(* Logix 5000 project; controller PLC_MCC1201_220AP1 vendor 1 type 14 code 164 rev 35.11; software revision 35.00 *) (continued)
   OSR_xStopCycle : BOOL;   // OSR stop cycle
   OS_xAreaSafetyOK : BOOL;   // OS area safety ok
   OS_xRequestAccessAreaOpSide : BOOL;   // OS access area request operator side
   OS_xRequestAccessAreaFarSide : BOOL;   // OS access area request far side
   OS_xConditionNotOKToCut : BOOL;   // OS condition not OK to cut
   OS_xConditionNotAllowedLower : BOOL;   // OS condition not allowed to lower head
   OS_xStopCycle : BOOL;   // OS stop cycle
   OS_xStartCycle : BOOL;   // OS start cycle
   OS_xDriveHomed : BOOL;   // OS drive homed
   AUX_tmOFF_DriveEnable : TIMER;   // Timer OFF retain drive enable
   AUX_tmOFF_AreaSafetyOK : TIMER;   // Timer OFF area safety OK
   AUX_tmON_FdbkError : TIMER;   // Timer ON feedback error
   AUX_tmON_TimeoutHome : TIMER;   // Timer ON timeout home
   AUX_tmON_TimeoutFW : TIMER;   // Timer ON timeout forward
   AUX_tmON_TimeoutBW : TIMER;   // Timer ON timeout backward
   AUX_tmOFF_LowerHeadNotAllowed : TIMER;   // Timer OFF Lower Head not allowed
   AUX_tmOFF_AdvanceTimeToRise : TIMER;   // Timer OFF Advance time to rise
   AUX_tmON_DelayTimeDescent : TIMER;   // Timer ON Delay time descent
   AUX_tmOFF_AdvanceTimeToLubrication : TIMER;   // Timer OFF Advance time to Lubrication
   AUX_tmON_DelayTimeLubrication : TIMER;   // Timer ON Delay time Lubrication
   AUX_tmON_TimeoutHeadPosition : TIMER;   // Timer ON head error position
   CONST_dHomePosition_cmm : DINT;   // Home position [mm/100]
   CONST_dAcceleration_m_s2 : DINT;   // Acceleration [m/s2]
   CONST_dDeceleration_m_s2 : DINT;   // Deceleration [m/s2]
END_STRUCT
END_TYPE

TYPE MAC_EMERGENCYXCUT_ALM :
STRUCT
   rgxStoppingFaults : DINT[2];   // Stopping faults
   rgxFaults : DINT[1];   // Faults
   rgxWarning : DINT[1];   // Warning
   rgdCodeAlarm : DINT[1];   // Code faults
END_STRUCT
END_TYPE

TYPE MAC_EMERGENCYXCUT_HMR :
STRUCT
   xMan_JogForwardFdbk : BOOL;   // Manual jog forward fdbk {x|x|x|x|O}
   xMan_JogBackwardFdbk : BOOL;   // Manual jog backward fdbk {x|x|x|x|O}
   xMan_DescentHeadFdbk : BOOL;   // Manual descent head fdbk {x|x|x|x|O}
   xMan_LubricationFdbk : BOOL;   // Manual lubrication fdbk {x|x|x|x|O}
   xMan_AirActivationFdbk : BOOL;   // Manual air activation fdbk {x|x|x|x|O}
   xCountinuousCuttingEnabled : BOOL;   // Countinuous cutting mode enabled {x|x|x|x|O}
   dMode : DINT;   // Machine mode (1=Manual 4=Automatic 7=Semiauto)
   dStatus : DINT;   // Machine status (1=Idle 3=Running 7=Anomaly)
   dZoneStatus : DINT;   // Zone status (1=CycleON 2=StopCycle 4=StartReq 8=StopReq)
   dDistanceFromSnaproll_cmm : DINT;   // Distance from snaproll [mm/100] {mm/100|mm|x|x|O}
   rHeadUsage_km : REAL;   // Head usage [km] {km|km|x|x|O}
END_STRUCT
END_TYPE

TYPE MAC_EMERGENCYXCUT_HMW :
STRUCT
   xMan_JogForward : BOOL;   // Manual jog forward {x|x|x|x|O}
   xMan_JogBackward : BOOL;   // Manual jog backward {x|x|x|x|O}
   xMan_DescentHead : BOOL;   // Manual descent head {x|x|x|x|O}
   xMan_Lubrication : BOOL;   // Manual lubrication {x|x|x|x|O}
   xMan_AirActivation : BOOL;   // Manual air activation {x|x|x|x|O}
   xResetHeadUsage : BOOL;   // Reset head usage {x|x|x|x|O}
   dLowerHeadDelayTime_ms : DINT;   // Lower head delay time [ms] {ms|s|0|3|O}
   dRiseHeadAdvanceTime_ms : DINT;   // Rise head advance time [ms] {ms|s|0|3|O}
   dOilRetainTime_ms : DINT;   // Oil retain time after rising [ms] {ms|s|-3|3|O}
   dOilAdvanceTime_ms : DINT;   // Oil advance time before lowering [ms] {ms|s|-3|3|O}
   dCulletStripeLength_cmm : DINT;   // Cullet stripe length [mm/100] {mm/100|mm|1000|6000|M}
   dDistanceFromSnaproll_cmm : DINT;   // Distance from snaproll [mm/100] {mm/100|mm|0|65000|M}
   xUpdateDistanceFromSnaproll : BOOL;   // Update distance from snaproll {x|x|x|x|M}
END_STRUCT
END_TYPE

TYPE MAC_EMERGENCYXCUT_IN_MOTION :
STRUCT
   DR_MAJ : MOTION_INSTRUCTION;   // Drive jog
   DR_MAM : MOTION_INSTRUCTION;   // Drive positioning
   DR_MAS : MOTION_INSTRUCTION;   // Drive stop
END_STRUCT
END_TYPE

TYPE MAC_EMERGENCYXCUT_OUT_MOTION :
STRUCT
   DR_MSO : MOTION_INSTRUCTION;   // Drive ON
   DR_MSF : MOTION_INSTRUCTION;   // Drive OFF
   DR_MASR : MOTION_INSTRUCTION;   // Drive reset faults
   DR_MAJ : MOTION_INSTRUCTION;   // Drive jog
   DR_MAM : MOTION_INSTRUCTION;   // Drive positioning
   DR_MCD : MOTION_INSTRUCTION;   // Drive change speed
   DR_MAS : MOTION_INSTRUCTION;   // Drive stop
   DR_MAH : MOTION_INSTRUCTION;   // Drive homing
END_STRUCT
END_TYPE

TYPE MAC_Zone_ML :
STRUCT
   ST_xSelManualMode : BOOL;   // Selection manual mode
   ST_xSelAutoMode : BOOL;   // Selection auto mode
   ST_xManualModeConditionOK : BOOL;   // Condition Ok for manual mode
   ST_xManuModeReq : BOOL;   // Manual mode request
   ST_xManualModeAccepted : BOOL;   // Manual mode accepted
   ST_xAutoModeAccepted : BOOL;   // Auto mode accepted
   ST_xConditionOKStopCycle : BOOL;   // Condition OK for stop cycle
   ST_xStartCycleRequest : BOOL;   // Start cycle request
   ST_xCycleON : BOOL;   // Cycle ON
   ST_xStopCycleRequest : BOOL;   // Stop cycle request
   ST_xStopCycleAccepted : BOOL;   // Stop cycle accepted
   ST_xStopCycleReqForFaults : BOOL;   // Stop cycle request for stopping faults
   ST_xStopCycleAcceptForFaults : BOOL;   // Stop cycle accepted for stopping faults
   ST_xStopCycleForSaturation : BOOL;   // Stop cycle for saturation on next zone and breaker not available
   ST_xConveyorsNotOK : BOOL;   // Conveyors not OK
   ST_xConditionOkPhaseAdvancement : BOOL;   // Condition OK phases advancement
   ST_xConditionOkCycleON : BOOL;   // Condition OK cycle ON
   ST_xCleaningConditionOK : BOOL;   // Cleaning condition OK
   ST_xReqCleaning : BOOL;   // Request cleaning
   ST_xCleaningAccepted : BOOL;   // Cleaning accepted
   ST_xReqCleaningByOperator : BOOL;   // Clean cycle request by operator
   ST_xEnableControlError : BOOL;   // Enable control error
   ST_xZoneError : BOOL;   // Zone error
   ST_xAlarmOff : BOOL;   // Alarm OFF
   ST_xConditionOkChangeSpeed : BOOL;   // Condition OK for change speed
   ST_xFaultsEnabled : BOOL;   // Faults Enabled
   ST_xReadyToReceiveGlass : BOOL;   // Zone ready to receive glass
   OSR_xStartCycle : BOOL;   // OSR Start cycle
   OSR_xStopCycle : BOOL;   // OSR Stop cycle
   OSR_xForceStopCycle : BOOL;   // OSR Force stop cycle
   OSR_xAlarmAcoustic : BOOL;   // OSR Alarm acoustic
   OSR_xAlarmMuting : BOOL;   // OSR Alarm muting
   OSR_xManualAccepted : BOOL;   // OSR Manual mode accepted
   OSR_xAutoAccepted : BOOL;   // OSR Auto mode accepted
   OS_xStartCycle : BOOL;   // OS Start cycle
   OS_xStopCycle : BOOL;   // OS Stop cycle
   OS_xForceStopCycle : BOOL;   // OS Force stop cycle
   OS_xAlarmAcoustic : BOOL;   // OS Alarm acoustic
   OS_xAlarmMuting : BOOL;   // OS Alarm muting
   OS_xManualAccepted : BOOL;   // OS Manual mode accepted
   OS_xAutoAccepted : BOOL;   // OS Auto mode accepted
   OS_xCleaningAccepted : BOOL;   // OS Cleaning Accepted
   INPUT_x24VdcVoltageON : BOOL;   // 24Vdc Voltage ON
   INPUT_xMainSwitch : BOOL;   // Main Switch
   INPUT_xMainEmergencyON : BOOL;   // Main Emergency ON
   INPUT_xUPSEmergencyON : BOOL;   // UPS Emergency ON
   INPUT_xAlarmSilence : BOOL;   // Alarm Silence Button
   INPUT_xAlarmReset : BOOL;   // Alarm Reset Button
   INPUT_xCulletAllow1 : BOOL;   // Cullet.Allow 1
   INPUT_xCulletAllow2 : BOOL;   // Cullet.Allow 2
   INPUT_xCulletAllow3 : BOOL;   // Cullet.Allow 3
   INPUT_xProtectionPowerSupplyConditioner1 : BOOL;   // Protection Power Supply Conditioner 1
   INPUT_xProtectionPowerSupplyConditioner2 : BOOL;   // Protection Power Supply Conditioner 2
   INPUT_xPowerFailure120V_Auxiliary1 : BOOL;   // Power failure supply 120Vac auxiliary 1
   INPUT_xPowerFailure120V_Auxiliary2 : BOOL;   // Power failure supply 120Vac auxiliary 2
   INPUT_xPowerSupplyOK : BOOL;   // Power supply OK
   INPUT_xPowerSupply24VLogic1 : BOOL;   // Power supply 24Vdc Logic 1
   INPUT_xPowerSupply24VLogic2 : BOOL;   // Power supply 24Vdc Logic 2
   INPUT_xPowerSupply24VLogic3 : BOOL;   // Power supply 24Vdc Logic 3
   INPUT_xPowerSupply24VLogic4 : BOOL;   // Power supply 24Vdc Logic 4
   INPUT_xPowerSupply24VDrive1 : BOOL;   // Power supply 24Vdc Drive 1
   INPUT_xPowerSupply24VDrive2 : BOOL;   // Power supply 24Vdc Drive 2
   INPUT_xPowerSupply480VDrive1 : BOOL;   // Alarm power supply 400/480Vac Drive 1
   INPUT_xPowerSupply480VDrive2 : BOOL;   // Alarm power supply 400/480Vac Drive 2
   INPUT_xEthernetSwitch24VON : BOOL;   // Ethernet Switch 24Vdc Voltage ON
   INPUT_xEthernetSwitchFault : BOOL;   // Ethernet Switch Fault
   INPUT_xEmergencyLocalization1 : BOOL;   // Emergency localization 1 A33SB1 Main Emergency Button MCC1201
   INPUT_xEmergencyLocalization2 : BOOL;   // Emergency localization 2 A34SB1 Main Emergency Button M203DROP OPERATOR SIDE
   INPUT_xEmergencyLocalization3 : BOOL;   // Emergency localization 3 A34SB2 Main Emergency Button M203DROP FAR SIDE
   INPUT_xEmergencyLocalization4 : BOOL;   // Emergency localization 4
   INPUT_xEmergencyLocalization5 : BOOL;   // Emergency localization 5
   INPUT_xEmergencyLocalization6 : BOOL;   // Emergency localization 6
   INPUT_xEmergencyLocalization7 : BOOL;   // Emergency localization 7
   INPUT_xEmergencyLocalization8 : BOOL;   // Emergency localization 7
   OUTPUT_xMainEmergencyLamp : BOOL;   // Main emergency ON
   OUTPUT_xUPSEmergencyLamp : BOOL;   // UPS emergency ON
   OUTPUT_xMCCSafetyLamp : BOOL;   // Safeties ON
   OUTPUT_xAcousticAlarm : BOOL;   // Acoustic alarm
   OUTPUT_xCulletAllow1 : BOOL;   // Cullet.Allow 1
   OUTPUT_xCulletAllow2 : BOOL;   // Cullet.Allow 2
   OUTPUT_xCulletAllow3 : BOOL;   // Cullet.Allow 3
   OUTPUT_xEmergencyLocalization1 : BOOL;   // Emergency localization 1
   OUTPUT_xEmergencyLocalization2 : BOOL;   // Emergency localization 2
   OUTPUT_xEmergencyLocalization3 : BOOL;   // Emergency localization 3
   OUTPUT_xEmergencyLocalization4 : BOOL;   // Emergency localization 4
   OUTPUT_xEmergencyLocalization5 : BOOL;   // Emergency localization 5
   OUTPUT_xEmergencyLocalization6 : BOOL;   // Emergency localization 6
   OUTPUT_xEmergencyLocalization7 : BOOL;   // Emergency localization 7
   AUX_dLehrSpeed_mm_min : DINT;   // Lehr speed [mm/min]
   AUX_dAutoSpeed_mm_min : DINT;   // Automatic speed [mm/min]
   AUX_dManualSpeed_mm_min : DINT;   // Manual speed [mm/min]
   tmON_ResetAlarm : TIMER;   // Reset alarm
   tmON_24Vdc : TIMER;   // Presence 24Vdc timer
   tmON_480Vca : TIMER;   // Presence 480Vca timer
   tmON_EmergencyOK : TIMER;   // Emergency OK timer
   tmON_Cycle : TIMER;   // Cycle ON timer
   tmON_ForceStop : TIMER;   // Force stop cycle timer
   tmON_CycleAcousticAlarm : TIMER;   // Cycle acoustic alarm timer
   tmON_ConveyorsNotOK : TIMER;   // Conveyors not ok
   AUX_tmOFF_ResetAlarm : TIMER;   // TOFF Reset alarm
END_STRUCT
END_TYPE

TYPE MAC_Zone_ML_ALM :
STRUCT
   rgxEmergency : DINT[1];   // Emergency
   rgxStoppingFault : DINT[1];   // Stopping faults
   rgxFault : DINT[1];   // Faults
   rgxWarning : DINT[1];   // Warning
   rgdFaultCode : DINT[1];   // Fault codes
END_STRUCT
END_TYPE

TYPE MAC_Zone_ML_HMR :
STRUCT
   xZoneAlarm : BOOL;   // Zone fault {x|x|x|x|O}
   xCleaningEnabled : BOOL;   // Cleaning enabled {x|x|x|x|O}
   dZoneMode : DINT;   // Zone mode (1=Manual 4=Automatic 8=Manual Req) {x|x|x|x|O}
   dZoneState : DINT;   // Zone status (1=CycleON 2=StopCyc 4=CycleReq 8=StopReq 1024=E-Stop) {x|x|x|x|O}
   dCabinetState : DINT;   // Cabinet status (0=OK; 1=General power alarm; 2=Local power alarm) {x|x|x|x|O}
   dCleaningState : DINT;   // Cleaning zone status (1=CycleON 2=StopCyc 4=CycleReq 8=StopReq) {x|x|x|x|O}
   dAutoSpeed_mm_min : DINT;   // Automatic speed [mm/min] {mm/min|m/min|x|x|O}
   dManualSpeed_mm_min : DINT;   // Manual speed [mm/min] {mm/min|m/min|x|x|O}
   dLehrSpeed_mm_min : DINT;   // Lehr speed [mm/min] {mm/min|m/min|x|x|O}
   rSpare : DINT;   // Spare
   rgxMan : DINT;   // Manual commands {x|x|x|x|O}
END_STRUCT
END_TYPE

TYPE MAC_Zone_ML_HMW :
STRUCT
   xManualModeReq : BOOL;   // Manual mode request {x|x|x|x|O}
   xAutoModeReq : BOOL;   // Automatic mode request {x|x|x|x|O}
   xStartCleanZoneRequest : BOOL;   // Start clean zone request {x|x|x|x|O}
   xStopCleanZoneRequest : BOOL;   // Stop clean zone request {x|x|x|x|O}
   xStartCycleRequest : BOOL;   // Start cycle request {x|x|x|x|O}
   xStopCycleRequest : BOOL;   // Stop cycle request {x|x|x|x|O}
   xForceStopCycle : BOOL;   // Force stop cycle {x|x|x|x|O}
   xResetErrorRequest : BOOL;   // Reset error request {x|x|x|x|O}
   dAutoSpeed_mm_min : DINT;   // Automatic speed [mm/min] {mm/min|m/min|7|90|O}
   dManualSpeed_mm_min : DINT;   // Manual speed [mm/min] {mm/min|m/min|2|20|O}
   rSpeedRatio : REAL;   // Speed ratio increment {%|%|0.0|2.0|O}
   rgxMan : DINT;   // Manual commands {x|x|x|x|O}
END_STRUCT
END_TYPE

TYPE STRUCT_AccessArea :
STRUCT
   tAccess : AOI_AccessArea_STRUCT[2];
   ST_xStopFault : BOOL;
   ST_xAccessAreaRequestInOneArea : BOOL;
   ST_xAccessAreaAcceptedInOneArea : BOOL;
   ST_xRequestResetPhase : BOOL;
END_STRUCT
END_TYPE

TYPE SYS_FaultRecord :
STRUCT
   TimeLow : DINT;
   TimeHigh : DINT;
   Type : INT;
   Code : INT;
   Info : DINT[8];
END_STRUCT
END_TYPE

TYPE UDT_CONSUMED_CULLET :   // Consumed tags from cullet system
STRUCT
   dSyncHead : DINT;   // Synchro head
   iCULLETtoMB_1 : INT;   // Status and Control
   iCULLETtoMB_2 : INT;   // Status and Control
   iCULLETtoMB_3 : INT;   // Spare
   iCULLETtoMB_4 : INT;   // Spare
   iCULLETtoMB_5 : INT;   // Spare
   iCULLETtoMB_6 : INT;   // Spare
   iCULLETtoMB_7 : INT;   // Spare
   iCULLETtoMB_8 : INT;   // Spare
   dSyncTail : DINT;   // Synchro tail
END_STRUCT
END_TYPE

TYPE UDT_CONSUMED_NEXT :   // Consumed tags from next section
STRUCT
   dSyncHead : DINT;   // Synchro head
   iM2toMB_1 : INT;   // Status and Control
   iM2toMB_2 : INT;   // Status and Control
   iM2toMB_3 : INT;   // Status and Control
   iM2toMB_4 : INT;   // Status and Control
   iM2toMB_5 : INT;   // Status and Control
   iM2toMB_6 : INT;   // Status and Control
   iM2toMB_7 : INT;   // Status and Control
   iM2toMB_8 : INT;   // Status and Control
   dSyncTail : DINT;   // Synchro tail
END_STRUCT
END_TYPE

TYPE UDT_MAN_CMD_WR :   // Manual commands from HMI
STRUCT
   CONV_Manual_ALL : BOOL;
   CONV_Man_ALL_FWD : BOOL;
   CONV_Man_ALL_REV : BOOL;
   M202M1_Manual : BOOL;
   M202M1_ManFWD : BOOL;
   M202M1_ManREV : BOOL;
   M202M1_ManSpeed : DINT;
   M202M1_TorqueIN : DINT;
   M203M1_Manual : BOOL;
   M203M1_ManFWD : BOOL;
   M203M1_ManREV : BOOL;
   M203M1_ManSpeed : DINT;
   M203M1_TorqueIN : DINT;
   M204M1_Manual : BOOL;
   M204M1_ManFWD : BOOL;
   M204M1_ManREV : BOOL;
   M204M1_ManSpeed : DINT;
   M204M1_TorqueIN : DINT;
   M206M1_Manual : BOOL;
   M206M1_ManFWD : BOOL;
   M206M1_ManREV : BOOL;
   M206M1_ManSpeed : DINT;
   M206M1_TorqueIN : DINT;
   M207M1_Manual : BOOL;
   M207M1_ManFWD : BOOL;
   M207M1_ManREV : BOOL;
   M207M1_ManSpeed : DINT;
   M207M1_TorqueIN : DINT;
   M208M1_Manual : BOOL;
   M208M1_ManFWD : BOOL;
   M208M1_ManREV : BOOL;
   M208M1_ManSpeed : DINT;
   M208M1_TorqueIN : DINT;
   M209M1_Manual : BOOL;
   M209M1_ManFWD : BOOL;
   M209M1_ManREV : BOOL;
   M209M1_ManSpeed : DINT;
   M209M1_TorqueIN : DINT;
   M210M1_Manual : BOOL;
   M210M1_ManFWD : BOOL;
   M210M1_ManREV : BOOL;
   M210M1_ManSpeed : DINT;
   M210M1_TorqueIN : DINT;
   M211M1_Manual : BOOL;
   M211M1_ManFWD : BOOL;
   M211M1_ManREV : BOOL;
   M211M1_ManSpeed : DINT;
   M211M1_TorqueIN : DINT;
   M212M1_Manual : BOOL;
   M212M1_ManFWD : BOOL;
   M212M1_ManREV : BOOL;
   M212M1_ManSpeed : DINT;
   M212M1_TorqueIN : DINT;
   M213M1_Manual : BOOL;
   M213M1_ManFWD : BOOL;
   M213M1_ManREV : BOOL;
   M213M1_ManSpeed : DINT;
   M213M1_TorqueIN : DINT;
   M213AM1_Manual : BOOL;
   M213AM1_ManFWD : BOOL;
   M213AM1_ManREV : BOOL;
   M213AM1_ManSpeed : DINT;
   M213AM1_TorqueIN : DINT;
   M213BM1_Manual : BOOL;
   M213BM1_ManFWD : BOOL;
   M213BM1_ManREV : BOOL;
   M213BM1_ManSpeed : DINT;
   M213BM1_TorqueIN : DINT;
   M214M1_Manual : BOOL;
   M214M1_ManFWD : BOOL;
   M214M1_ManREV : BOOL;
   M214M1_ManSpeed : DINT;
   M214M1_TorqueIN : DINT;
   M215M1_Manual : BOOL;
   M215M1_ManFWD : BOOL;
   M215M1_ManREV : BOOL;
   M215M1_ManSpeed : DINT;
   M215M1_TorqueIN : DINT;
   M216M1_Manual : BOOL;
   M216M1_ManFWD : BOOL;
   M216M1_ManREV : BOOL;
   M216M1_ManSpeed : DINT;
   M216M1_TorqueIN : DINT;
   M217M1_Manual : BOOL;
   M217M1_ManFWD : BOOL;
   M217M1_ManREV : BOOL;
   M217M1_ManSpeed : DINT;
   M217M1_TorqueIN : DINT;
   M218M1_Manual : BOOL;
   M218M1_ManFWD : BOOL;
   M218M1_ManREV : BOOL;
   M218M1_ManSpeed : DINT;
   M218M1_TorqueIN : DINT;
   M219M1_Manual : BOOL;
   M219M1_ManFWD : BOOL;
   M219M1_ManREV : BOOL;
   M219M1_ManSpeed : DINT;
   M219M1_TorqueIN : DINT;
   M220M1_Manual : BOOL;
   M220M1_ManFWD : BOOL;
   M220M1_ManREV : BOOL;
   M220M1_ManSpeed : DINT;
   M220M1_TorqueIN : DINT;
   M225M1_Manual : BOOL;
   M225M1_ManFWD : BOOL;
   M225M1_ManREV : BOOL;
   M225M1_ManSpeed : DINT;
   M225M1_TorqueIN : DINT;
   M301M1_Manual : BOOL;
   M301M1_ManFWD : BOOL;
   M301M1_ManREV : BOOL;
   M301M1_ManSpeed : DINT;
   M301M1_TorqueIN : DINT;
   M301M2_Manual : BOOL;
   M301M2_ManFWD : BOOL;
   M301M2_ManREV : BOOL;
   M301M2_ManSpeed : DINT;
   M301M2_TorqueIN : DINT;
END_STRUCT
END_TYPE

TYPE UDT_MOTOR_HMR :
STRUCT
   M202M1_Feedback : BOOL;
   M202M1_Faulted : BOOL;
   M202M1_FaultCode : DINT;
   M202M1_OutSpeed : DINT;
   M202M1_OutCurrent : DINT;
   M202M1_OutTorque : DINT;
   M203M1_Feedback : BOOL;
   M203M1_Faulted : BOOL;
   M203M1_FaultCode : DINT;
   M203M1_OutSpeed : DINT;
   M203M1_OutCurrent : DINT;
   M203M1_OutTorque : DINT;
   M204M1_Feedback : BOOL;
   M204M1_Faulted : BOOL;
   M204M1_FaultCode : DINT;
   M204M1_OutSpeed : DINT;
   M204M1_OutCurrent : DINT;
   M205M1_Feedback : BOOL;
   M205M1_Faulted : BOOL;
   M205M1_FaultCode : DINT;
   M205M1_OutSpeed : DINT;
   M205M1_OutCurrent : DINT;
   M205M1_OutTorque : DINT;
   M206M1_Feedback : BOOL;
   M206M1_Faulted : BOOL;
   M206M1_FaultCode : DINT;
   M206M1_OutSpeed : DINT;
   M206M1_OutCurrent : DINT;
   M206M1_OutTorque : DINT;
   M207M1_Feedback : BOOL;
   M207M1_Faulted : BOOL;
   M207M1_FaultCode : DINT;
   M207M1_OutSpeed : DINT;
   M207M1_OutCurrent : DINT;
   M207M1_OutTorque : DINT;
   M208M1_Feedback : BOOL;
   M208M1_Faulted : BOOL;
   M208M1_FaultCode : DINT;
   M208M1_OutSpeed : DINT;
   M208M1_OutCurrent : DINT;
   M208M1_OutTorque : DINT;
   M209M1_Feedback : BOOL;
   M209M1_Faulted : BOOL;
   M209M1_FaultCode : DINT;
   M209M1_OutSpeed : DINT;
   M209M1_OutCurrent : DINT;
   M209M1_OutTorque : DINT;
   M210M1_Feedback : BOOL;
   M210M1_Faulted : BOOL;
   M210M1_FaultCode : DINT;
   M210M1_OutSpeed : DINT;
   M210M1_OutCurrent : DINT;
   M210M1_OutTorque : DINT;
   M211M1_Feedback : BOOL;
   M211M1_Faulted : BOOL;
   M211M1_FaultCode : DINT;
   M211M1_OutSpeed : DINT;
   M211M1_OutCurrent : DINT;
   M211M1_OutTorque : DINT;
   M212M1_Feedback : BOOL;
   M212M1_Faulted : BOOL;
   M212M1_FaultCode : DINT;
   M212M1_OutSpeed : DINT;
   M212M1_OutCurrent : DINT;
   M212M1_OutTorque : DINT;
   M213M1_Feedback : BOOL;
   M213M1_Faulted : BOOL;
   M213M1_FaultCode : DINT;
   M213M1_OutSpeed : DINT;
   M213M1_OutCurrent : DINT;
   M213M1_OutTorque : DINT;
   M213AM1_Feedback : BOOL;
   M213AM1_Faulted : BOOL;
   M213AM1_FaultCode : DINT;
   M213AM1_OutSpeed : DINT;
   M213AM1_OutCurrent : DINT;
   M213AM1_OutTorque : DINT;
   M213BM1_Feedback : BOOL;
   M213BM1_Faulted : BOOL;
   M213BM1_FaultCode : DINT;
   M213BM1_OutSpeed : DINT;
   M213BM1_OutCurrent : DINT;
   M213BM1_OutTorque : DINT;
   M214M1_Feedback : BOOL;
   M214M1_Faulted : BOOL;
   M214M1_FaultCode : DINT;
   M214M1_OutSpeed : DINT;
   M214M1_OutCurrent : DINT;
   M214M1_OutTorque : DINT;
   M215M1_Feedback : BOOL;
   M215M1_Faulted : BOOL;
   M215M1_FaultCode : DINT;
   M215M1_OutSpeed : DINT;
   M215M1_OutCurrent : DINT;
   M215M1_OutTorque : DINT;
   M216M1_Feedback : BOOL;
   M216M1_Faulted : BOOL;
   M216M1_FaultCode : DINT;
   M216M1_OutSpeed : DINT;
   M216M1_OutCurrent : DINT;
   M216M1_OutTorque : DINT;
   M217M1_Feedback : BOOL;
   M217M1_Faulted : BOOL;
   M217M1_FaultCode : DINT;
   M217M1_OutSpeed : DINT;
   M217M1_OutCurrent : DINT;
   M217M1_OutTorque : DINT;
   M218M1_Feedback : BOOL;
   M218M1_Faulted : BOOL;
   M218M1_FaultCode : DINT;
   M218M1_OutSpeed : DINT;
   M218M1_OutCurrent : DINT;
   M218M1_OutTorque : DINT;
   M219M1_Feedback : BOOL;
   M219M1_Faulted : BOOL;
   M219M1_FaultCode : DINT;
   M219M1_OutSpeed : DINT;
   M219M1_OutCurrent : DINT;
   M219M1_OutTorque : DINT;
   M220M1_Feedback : BOOL;
   M220M1_Faulted : BOOL;
   M220M1_FaultCode : DINT;
   M220M1_OutSpeed : DINT;
   M220M1_OutCurrent : DINT;
   M220M1_OutTorque : DINT;
   M225M1_Feedback : BOOL;
   M225M1_Faulted : BOOL;
   M225M1_FaultCode : DINT;
   M225M1_OutSpeed : DINT;
   M225M1_OutCurrent : DINT;
   M225M1_OutTorque : DINT;
   M301M1_Feedback : BOOL;
   M301M1_Faulted : BOOL;
   M301M1_FaultCode : DINT;
   M301M1_OutSpeed : DINT;
   M301M1_OutCurrent : DINT;
   M301M1_OutTorque : DINT;
   M301M2_Feedback : BOOL;
   M301M2_Faulted : BOOL;
   M301M2_FaultCode : DINT;
   M301M2_OutSpeed : DINT;
   M301M2_OutCurrent : DINT;
   M301M2_OutTorque : DINT;
END_STRUCT
END_TYPE

TYPE UDT_PRODUCED_CULLET :   // Produced tags for cullet system
STRUCT
   dSyncHead : DINT;   // Synchro head
   MBtoCULLET_1 : INT;   // Status and Control
   MBtoCULLET_2 : INT;   // Status and Control
   MBtoCULLET_3 : INT;   // Status and Control
   MBtoCULLET_4 : INT;   // Status and Control
   MBtoCULLET_5 : INT;   // Status and Control
   MBtoCULLET_6 : INT;   // Status and Control
   MBtoCULLET_7 : INT;   // Status and Control
   MBtoCULLET_8 : INT;   // Status and Control
   dSyncTail : DINT;   // Synchro tail
END_STRUCT
END_TYPE

TYPE UDT_PRODUCED_NEXT :   // Produced tags for next section
STRUCT
   dSyncHead : DINT;   // Synchro head
   iMBtoM2_1 : INT;   // Spare
   iMBtoM2_2 : INT;   // Lehr Speed [IPM x 10]
   iMBtoM2_3 : INT;   // Status and Control
   iMBtoM2_4 : INT;   // Status and Control
   iMBtoM2_5 : INT;   // Status and Control
   iMBtoM2_6 : INT;   // Spare
   iMBtoM2_7 : INT;   // Spare
   iMBtoM2_8 : INT;   // Spare
   dSyncTail : DINT;   // Synchro tail
END_STRUCT
END_TYPE

TYPE UDT_Spare32bit_Alm :   // Generic base Structure for Fault, alarm and warning
STRUCT
   x0 : BOOL;   // Spare 0
   x1 : BOOL;   // Spare 1
   x2 : BOOL;   // Spare 2
   x3 : BOOL;   // Spare 3
   x4 : BOOL;   // Spare 4
   x5 : BOOL;   // Spare 5
   x6 : BOOL;   // Spare 6
   x7 : BOOL;   // Spare 7
   x8 : BOOL;   // Spare 8
   x9 : BOOL;   // Spare 9
   x10 : BOOL;   // Spare 10
   x11 : BOOL;   // Spare 11
   x12 : BOOL;   // Spare 12
   x13 : BOOL;   // Spare 13
   x14 : BOOL;   // Spare 14
   x15 : BOOL;   // Spare 15
   x16 : BOOL;   // Spare 16
   x17 : BOOL;   // Spare 17
   x18 : BOOL;   // Spare 18
   x19 : BOOL;   // Spare 19
   x20 : BOOL;   // Spare 20
   x21 : BOOL;   // Spare 21
   x22 : BOOL;   // Spare 22
   x23 : BOOL;   // Spare 23
   x24 : BOOL;   // Spare 24
   x25 : BOOL;   // Spare 25
   x26 : BOOL;   // Spare 26
   x27 : BOOL;   // Spare 27
   x28 : BOOL;   // Spare 28
   x29 : BOOL;   // Spare 29
   x30 : BOOL;   // Spare 30
   x31 : BOOL;   // Spare 31
END_STRUCT
END_TYPE

TYPE ZONE_UPS :
STRUCT
   ST_xZoneError : BOOL;   // Zone error
   ST_xSelectionAutoMode : BOOL; {access None}   // Automatic mode selection
   ST_xSelectionManualMode : BOOL; {access None}   // Manual mode selection
   ST_xConditionOKManualMode : BOOL; {access None}   // Condition OK for manual mode
   ST_xManualModeAccepted : BOOL; {access None}   // Manual mode accepted
   ST_xAutoModeAccepted : BOOL; {access None}   // Automatic mode accepted
   ST_xManualModeRequest : BOOL; {access None}   // Manual mode request
   ST_xFaultsEnabled : BOOL;   // Faults enabled
   ST_xZoneEmergency : BOOL;   // Cumulative of emergency faults active
   ST_xZoneFaults : BOOL;   // Cumulative of zone faults
   ST_xZoneStoppingFaults : BOOL;   // Cumulative of zone stopping faults
   ST_xZoneWarnings : BOOL;   // Cumulative of zone warning
   ST_xConditionOKStopCycle : BOOL;   // Condition OK for stop cycle
   ST_xStartCycleRequest : BOOL;   // Start cycle request
   ST_xCycleON : BOOL;   // Cycle ON
   ST_xStopCycleRequest : BOOL;   // Stop cycle request
   ST_xStopCycleAccepted : BOOL;   // Stop cycle accepted
   ST_xStopCycleReqForFaults : BOOL;   // Stop cycle request for stopping faults
   ST_xStopCycleAcceptForFaults : BOOL;   // Stop cycle accepted for stopping faults
   ST_xConditionOkPhaseAdvancement : BOOL;   // Condition OK phases advancement
   ST_xConditionOkCycleON : BOOL;   // Condition OK cycle ON
   OSR_xStartCycle : BOOL;   // OSR Start cycle
   OSR_xStopCycle : BOOL;   // OSR Stop cycle
   OSR_xForceStopCycle : BOOL;   // OSR Force stop cycle
   OS_xStartCycle : BOOL;   // OS Start cycle
   OS_xStopCycle : BOOL;   // OS Stop cycle
   OS_xForceStopCycle : BOOL;   // OS Force stop cycle
   INPUT_x24vdcVoltageOn : BOOL;   // INPUT.L+.24VDC Voltage ON
   INPUT_xPowerFailurePLCA : BOOL;   // INPUT.QF.Power failure PLC A
   INPUT_xPowerFailurePLCB : BOOL;   // INPUT.QF.Power failure PLC B
   INPUT_xUPSEmergencyON : BOOL;   // INPUT.KE.UPS Emergency ON
   INPUT_xEmLocUps1 : BOOL;   // INPUT.A33SB2.Emergency localization UPS 203DROP OPERATOR SIDE
   INPUT_xEmLocUps2 : BOOL;   // INPUT.A33SB3.Emergency localization UPS 203DROP FAR SIDE
   INPUT_xEmLocUps3 : BOOL;   // INPUT.A33SB4.Emergency localization UPS M225 FAR SIDE
   INPUT_xEmLocUps4 : BOOL;   // INPUT.A33SB5.Emergency localization UPS CS4225
   INPUT_xEmLocUps5 : BOOL;   // INPUT.Emergency localization UPS
   INPUT_xEmLocUps6 : BOOL;   // INPUT.Emergency localization UPS
   INPUT_xEmLocUps7 : BOOL;   // INPUT.Emergency localization UPS
   INPUT_xEmLocUps8 : BOOL;   // INPUT.Emergency localization UPS
   INPUT_xClutchON : BOOL;   // INPUT.Clutch ON
   INPUT_xClutchOFF : BOOL;   // INPUT.Clutch OFF
   INPUT_xM200ClutchON : BOOL;   // INPUT.M200 Clutch ON
   INPUT_xM202ClutchON : BOOL;   // INPUT.M202 Clutch ON
   OUTPUT_xEmergencyUPSOn : BOOL;   // OUTPUT.HL.Emergency UPS On
   AUX_tmOFF_ResetAlarm : TIMER;   // Reset alarm
   AUX_tmON_24Vdc : TIMER;   // Presence 24Vdc timer
   AUX_tmON_EmergencyOK : TIMER;   // Emergency OK timer
   AUX_tmON_Clutch1feedback : TIMER;   // Feedback error clutch
   AUX_tmON_Clutch2feedback : TIMER;   // Feedback error clutch
END_STRUCT
END_TYPE

TYPE ZONE_UPS_ALM :
STRUCT
   rgxEmergency : DINT[1];   // Emergency alarms
   rgxStoppingFaults : DINT[2];   // Stopping faults
   rgxFaults : DINT[1];   // Faults
   rgxWarning : DINT[1];   // Warning
   rgdCodeAlarm : DINT[1];   // Code faults
END_STRUCT
END_TYPE

TYPE ZONE_UPS_HMR :
STRUCT
   dZoneMode : DINT;   // Zone modality (1=Manual;4=Automatic;8=Manual request) {x|x|x|x|O}
   xZoneAlarm : BOOL;   // Zone alarm {x|x|x|x|O}
   dZoneState : DINT;   // Zone status (1=CycleON 2=StopCyc 4=CycleReq 8=StopReq 1024=E-Stop) {x|x|x|x|O}
END_STRUCT
END_TYPE

TYPE ZONE_UPS_HMW :
STRUCT
   xResetErrorRequest : BOOL;   // Reset error request {x|x|x|x|O}
   xAutoModeReq : BOOL;   // Automatic mode request {x|x|x|x|O}
   xManModeReq : BOOL;   // Manual mode request {x|x|x|x|O}
   xStartCycleRequest : BOOL;   // Start cycle request {x|x|x|x|O}
   xStopCycleRequest : BOOL;   // Stop cycle request {x|x|x|x|O}
   xForceStopCycle : BOOL;   // Force stop cycle {x|x|x|x|O}
END_STRUCT
END_TYPE

ADD_ON_INSTRUCTION AOI_AccessArea   (* revision 1.0 *)
VAR_INPUT
   IN_xConditionOkForce : BOOL; {access None, required}
   IN_xConditionOkForAccess : BOOL; {access None, required}
   IN_xAccButton : BOOL; {access None, required}
   IN_xAccSelector : BOOL; {access None, required}
   IN_xLampClock : BOOL; {access None, required}
END_VAR
VAR_OUTPUT
   OUT_xOpeningDoor : BOOL; {access None, required}
   OUT_xLamp : BOOL; {access None, required}
   OUT_xAccessRequest : BOOL; {access None}
   OUT_xAccessAccepted : BOOL; {access None}
END_VAR
VAR
   tSTC : AOI_AccessArea_GP_STC; {access None}
END_VAR

ROUTINE Logic   (* ladder *)
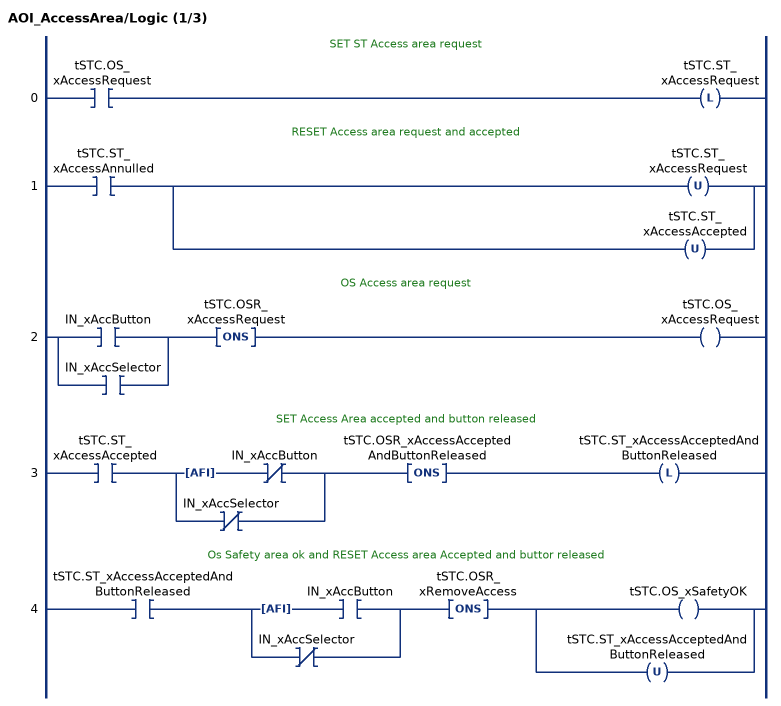
   // SET ST Access area request
   0: XIC(tSTC.OS_xAccessRequest)OTL(tSTC.ST_xAccessRequest);
   // RESET Access area request and accepted
   1: XIC(tSTC.ST_xAccessAnnulled)[OTU(tSTC.ST_xAccessRequest) ,OTU(tSTC.ST_xAccessAccepted) ];
   // OS Access area request
   2: [XIC(IN_xAccButton) ,XIC(IN_xAccSelector) ]ONS(tSTC.OSR_xAccessRequest)OTE(tSTC.OS_xAccessRequest);
   // SET Access Area accepted and button released
   3: XIC(tSTC.ST_xAccessAccepted)[AFI() XIO(IN_xAccButton) ,XIO(IN_xAccSelector) ]ONS(tSTC.OSR_xAccessAcceptedAndButtonReleased)OTL(tSTC.ST_xAccessAcceptedAndButtonReleased);
   // Os Safety area ok and RESET Access area Accepted and buttor released
   4: XIC(tSTC.ST_xAccessAcceptedAndButtonReleased)[AFI() XIC(IN_xAccButton) ,XIO(IN_xAccSelector) ]ONS(tSTC.OSR_xRemoveAccess)[OTE(tSTC.OS_xSafetyOK) ,OTU(tSTC.ST_xAccessAcceptedAndButtonReleased) ];
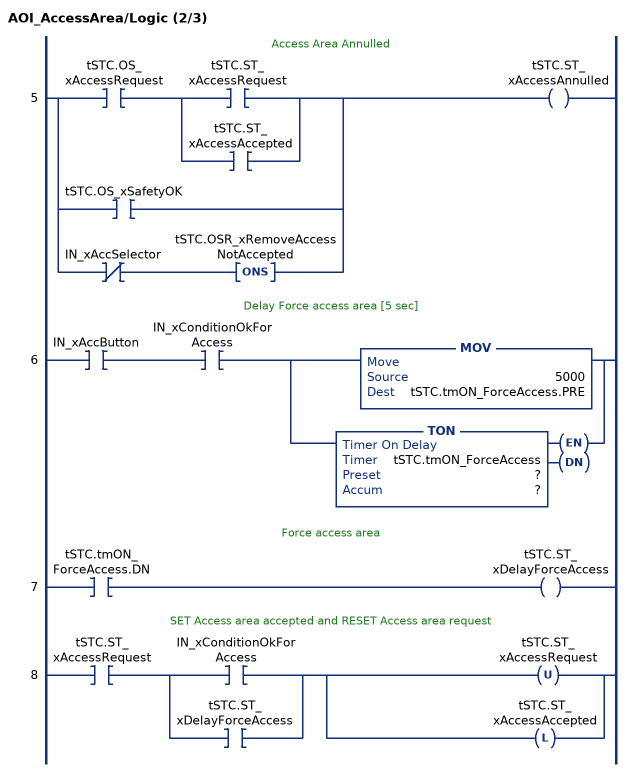
   // Access Area Annulled
   5: [XIC(tSTC.OS_xAccessRequest) [XIC(tSTC.ST_xAccessRequest) ,XIC(tSTC.ST_xAccessAccepted) ] ,XIC(tSTC.OS_xSafetyOK) ,XIO(IN_xAccSelector) ONS(tSTC.OSR_xRemoveAccessNotAccepted) ]OTE(tSTC.ST_xAccessAnnulled);
   // Delay Force access area [5 sec]
   6: XIC(IN_xAccButton)XIC(IN_xConditionOkForAccess)[MOV(5000,tSTC.tmON_ForceAccess.PRE) ,TON(tSTC.tmON_ForceAccess,?,?) ];
   // Force access area
   7: XIC(tSTC.tmON_ForceAccess.DN)OTE(tSTC.ST_xDelayForceAccess);
   // SET Access area accepted and RESET Access area request
   8: XIC(tSTC.ST_xAccessRequest)[XIC(IN_xConditionOkForAccess) ,XIC(tSTC.ST_xDelayForceAccess) ][OTU(tSTC.ST_xAccessRequest) ,OTL(tSTC.ST_xAccessAccepted) ];
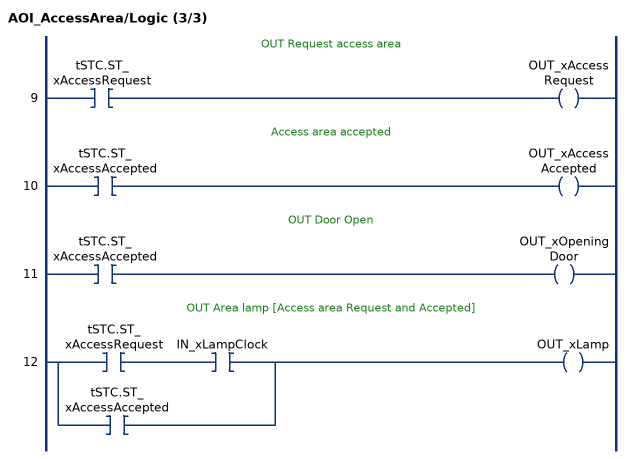
   // OUT Request access area
   9: XIC(tSTC.ST_xAccessRequest)OTE(OUT_xAccessRequest);
   // Access area accepted
   10: XIC(tSTC.ST_xAccessAccepted)OTE(OUT_xAccessAccepted);
   // OUT Door Open
   11: XIC(tSTC.ST_xAccessAccepted)OTE(OUT_xOpeningDoor);
   // OUT Area lamp [Access area Request and Accepted]
   12: [XIC(tSTC.ST_xAccessRequest) XIC(IN_xLampClock) ,XIC(tSTC.ST_xAccessAccepted) ]OTE(OUT_xLamp);
END_ROUTINE
END_ADD_ON_INSTRUCTION
